// TIA Portal project "TIA1200_Level1" (V19) (continued)
REGION Network 5: Retract Cylinder B logic
   // Retract cylinder B after both cylinders are extended
   RUNG wire#powerrail
      Contact( "Gripper open" )
      Contact( "Cylinder A extended" )
      Contact( "Cylinder B extended" )
      S_SR(operand := "Retract cylinder B", r1 := wire#w1)
   END_RUNG
   RUNG wire#powerrail
      Contact( "Cylinder B retracted" )
   END_RUNG wire#w1
   // the same network as SCL:
   IF "Gripper open" AND "Cylinder A extended" AND "Cylinder B extended" THEN
       "Retract cylinder B" := TRUE;   // SR flip-flop
   END_IF;
   IF "Cylinder B retracted" THEN "Retract cylinder B" := FALSE; END_IF;
END_REGION

REGION Network 6: Retract Cylinder A Logic
   // Retract cylinder A when cylinder A is extended, cylinder B is retracted and gripper is open; stop after its upper limit
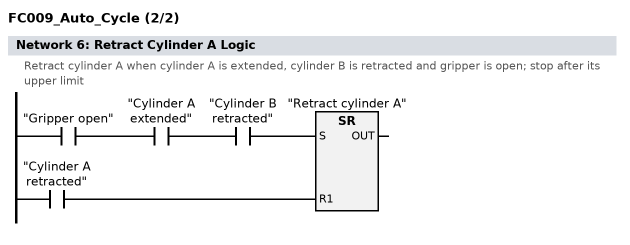
   RUNG wire#powerrail
      Contact( "Gripper open" )
      Contact( "Cylinder A extended" )
      Contact( "Cylinder B retracted" )
      S_SR(operand := "Retract cylinder A", r1 := wire#w1)
   END_RUNG
   RUNG wire#powerrail
      Contact( "Cylinder A retracted" )
   END_RUNG wire#w1
   // the same network as SCL:
   IF "Gripper open" AND "Cylinder A extended" AND "Cylinder B retracted" THEN
       "Retract cylinder A" := TRUE;   // SR flip-flop
   END_IF;
   IF "Cylinder A retracted" THEN "Retract cylinder A" := FALSE; END_IF;
END_REGION
END_FUNCTION

FUNCTION "FC010_OneButton_OneLight" : Void   // FC14, LAD
{ S7_Optimized_Access := 'TRUE' }
VERSION : 0.1
   VAR_TEMP   // added for the SCL form of the ladder/FBD networks
      _w1 : Bool;
   END_VAR
BEGIN

REGION Network 1 (FBD): Lamp Toggle Logic
   // XOR outputs 1 only when both inputs have different states; identical states produce 0
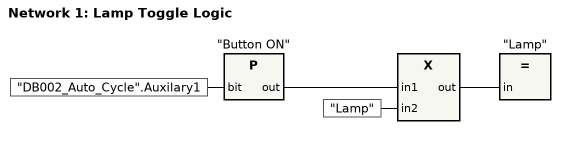
   #_w1 := "Button ON" AND NOT "DB002_Auto_Cycle".Auxilary1;   // rising edge of "Button ON"
   "DB002_Auto_Cycle".Auxilary1 := "Button ON";
   "Lamp" := #_w1 XOR "Lamp";
END_REGION
END_FUNCTION

FUNCTION "FC011_Voltage_Control" : Void   // FC15, LAD
{ S7_Optimized_Access := 'TRUE' }
VERSION : 0.1
BEGIN

REGION Network 1: Voltage Output Control Logic
   // Set QW80 to 0 V, 5 V, or 10 V depending on input states I1.0 and I1.1 (Integer range: 0 - 27648)
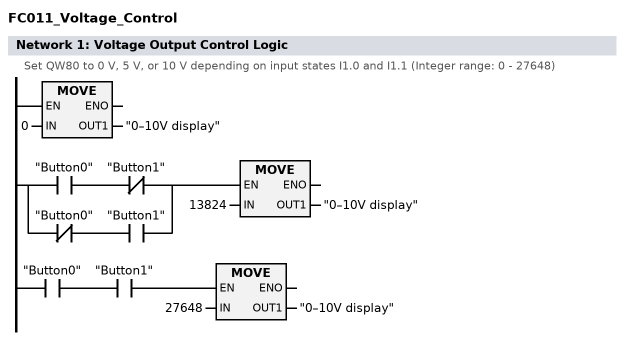
   RUNG wire#powerrail
      Move(in := 0, out1 => "0–10V display")
   END_RUNG
   RUNG wire#powerrail
      Contact( "Button0" )
      I_Contact( "Button1" )
      wire#w1
      Move(in := 13824, out1 => "0–10V display")
   END_RUNG
   RUNG wire#powerrail
      I_Contact( "Button0" )
      Contact( "Button1" )
   END_RUNG wire#w1
   RUNG wire#powerrail
      Contact( "Button0" )
      Contact( "Button1" )
      Move(in := 27648, out1 => "0–10V display")
   END_RUNG
   // the same network as SCL:
   "0–10V display" := 0;
   IF ("Button0" AND NOT "Button1") OR (NOT "Button0" AND "Button1") THEN "0–10V display" := 13824; END_IF;
   IF "Button0" AND "Button1" THEN "0–10V display" := 27648; END_IF;
END_REGION
END_FUNCTION

FUNCTION "FC012_Calculations" : Void   // FC16, LAD
{ S7_Optimized_Access := 'TRUE' }
VERSION : 0.1
   VAR_TEMP   // added for the SCL form of the ladder/FBD networks
      _w1 : Bool;
   END_VAR
BEGIN

REGION Network 1: Production Stock Calculation
   // Calculate stock = Sum1 + Sum2 − Losses
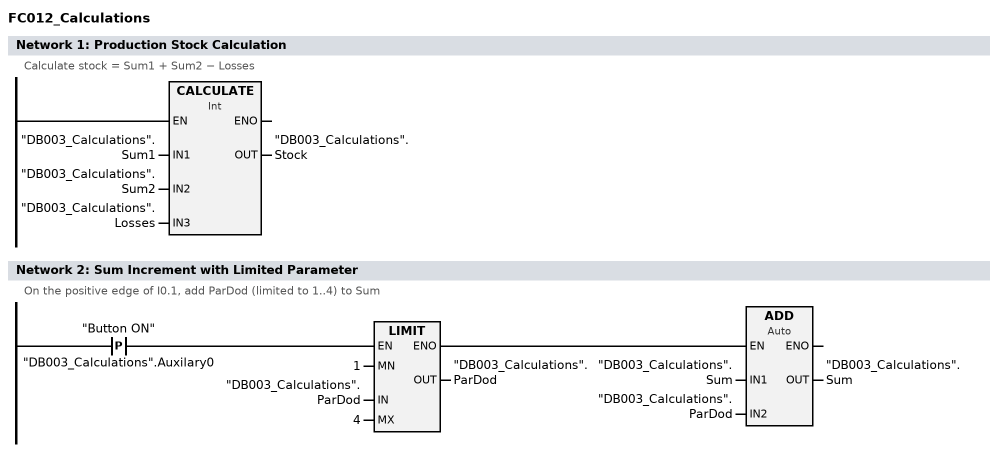
   RUNG wire#powerrail
      { S7_Templates := "SrcType := Int"; S7_Expression := "IN1 + IN2 - IN3" } Calculate(in1 := "DB003_Calculations".Sum1, in2 := "DB003_Calculations".Sum2, in3 := "DB003_Calculations".Losses, out => "DB003_Calculations".Stock)
   END_RUNG
   // the same network as SCL:
   "DB003_Calculations".Stock := "DB003_Calculations".Sum1 + "DB003_Calculations".Sum2 - "DB003_Calculations".Losses;
END_REGION

REGION Network 2: Sum Increment with Limited Parameter
   // On the positive edge of I0.1, add ParDod (limited to 1..4) to Sum
   #_w1 := "Button ON" AND NOT "DB003_Calculations".Auxilary0;   // rising edge of "Button ON"
   "DB003_Calculations".Auxilary0 := "Button ON";
   IF #_w1 THEN
       "DB003_Calculations".ParDod := LIMIT(MN := 1, IN := "DB003_Calculations".ParDod, MX := 4);
       "DB003_Calculations".Sum := "DB003_Calculations".Sum + "DB003_Calculations".ParDod;
   END_IF;
END_REGION
END_FUNCTION

FUNCTION "FC013_Labeler_Control" : Void   // FC17, LAD
{ S7_Optimized_Access := 'TRUE' }
VERSION : 0.1
   VAR_TEMP   // added for the SCL form of the ladder/FBD networks
      _w1 : Bool;
   END_VAR
BEGIN

REGION Network 1: Roll Initialization & Roll Counter
   // On Button0 load a new labels roll and increment labels roll total counter
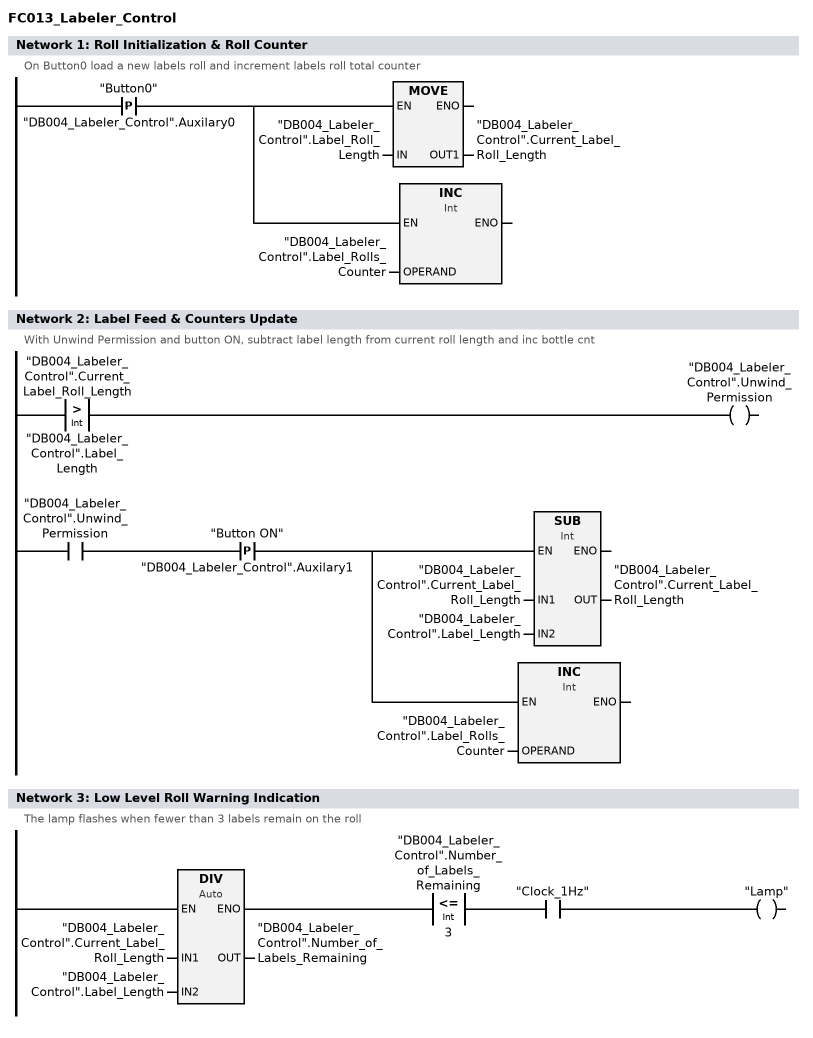
   RUNG wire#powerrail
      P_Contact(operand := "Button0", bit := "DB004_Labeler_Control".Auxilary0)
      wire#w1
      Move(in := "DB004_Labeler_Control".Label_Roll_Length, out1 => "DB004_Labeler_Control".Current_Label_Roll_Length)
   END_RUNG
   RUNG wire#w1
      { S7_Templates := "DestType := Int" } Inc( "DB004_Labeler_Control".Label_Rolls_Counter )
   END_RUNG
   // the same network as SCL:
   #_w1 := "Button0" AND NOT "DB004_Labeler_Control".Auxilary0;   // rising edge of "Button0"
   "DB004_Labeler_Control".Auxilary0 := "Button0";
   IF #_w1 THEN
       "DB004_Labeler_Control".Current_Label_Roll_Length := "DB004_Labeler_Control".Label_Roll_Length;
       "DB004_Labeler_Control".Label_Rolls_Counter := "DB004_Labeler_Control".Label_Rolls_Counter + 1;
   END_IF;
END_REGION

REGION Network 2: Label Feed & Counters Update
   // With Unwind Permission and button ON, subtract label length from current roll length and inc bottle cnt
   RUNG wire#powerrail
      { S7_Templates := "SrcType := Int" } GT_Contact(in1 := "DB004_Labeler_Control".Current_Label_Roll_Length, in2 := "DB004_Labeler_Control".Label_Length)
      Coil( "DB004_Labeler_Control".Unwind_Permission )
   END_RUNG
   RUNG wire#powerrail
      Contact( "DB004_Labeler_Control".Unwind_Permission )
      P_Contact(operand := "Button ON", bit := "DB004_Labeler_Control".Auxilary1)
      wire#w1
      { S7_Templates := "SrcType := Int" } Sub(in1 := "DB004_Labeler_Control".Current_Label_Roll_Length, in2 := "DB004_Labeler_Control".Label_Length, out => "DB004_Labeler_Control".Current_Label_Roll_Length)
   END_RUNG
   RUNG wire#w1
      { S7_Templates := "DestType := Int" } Inc( "DB004_Labeler_Control".Label_Rolls_Counter )
   END_RUNG
   // the same network as SCL:
   "DB004_Labeler_Control".Unwind_Permission := "DB004_Labeler_Control".Current_Label_Roll_Length > "DB004_Labeler_Control".Label_Length;
   #_w1 := "DB004_Labeler_Control".Unwind_Permission AND "Button ON" AND NOT "DB004_Labeler_Control".Auxilary1;   // rising edge of "Button ON"
   "DB004_Labeler_Control".Auxilary1 := "Button ON";
   IF #_w1 THEN
       "DB004_Labeler_Control".Current_Label_Roll_Length := "DB004_Labeler_Control".Current_Label_Roll_Length - "DB004_Labeler_Control".Label_Length;
       "DB004_Labeler_Control".Label_Rolls_Counter := "DB004_Labeler_Control".Label_Rolls_Counter + 1;
   END_IF;
END_REGION

REGION Network 3: Low Level Roll Warning Indication
   // The lamp flashes when fewer than 3 labels remain on the roll
   RUNG wire#powerrail
      Div(in1 := "DB004_Labeler_Control".Current_Label_Roll_Length, in2 := "DB004_Labeler_Control".Label_Length, out => "DB004_Labeler_Control".Number_of_Labels_Remaining)
      { S7_Templates := "SrcType := Int" } LE_Contact(in1 := "DB004_Labeler_Control".Number_of_Labels_Remaining, in2 := 3)
      Contact( "Clock_1Hz" )
      Coil( "Lamp" )
   END_RUNG
   // the same network as SCL:
   "DB004_Labeler_Control".Number_of_Labels_Remaining := "DB004_Labeler_Control".Current_Label_Roll_Length / "DB004_Labeler_Control".Label_Length;
   "Lamp" := ("DB004_Labeler_Control".Number_of_Labels_Remaining <= 3) AND "Clock_1Hz";
END_REGION
END_FUNCTION

FUNCTION "FC014_Buffer_Filling" : Void   // FC18, LAD
{ S7_Optimized_Access := 'TRUE' }
VERSION : 0.1
BEGIN

REGION Network 1: Buffer Counter & Limits Logic
   // Count up on I1.3 and down on I1.5 with CTUD (PV=10). NOT QU blocks further up-counting at full; reset with I0.0
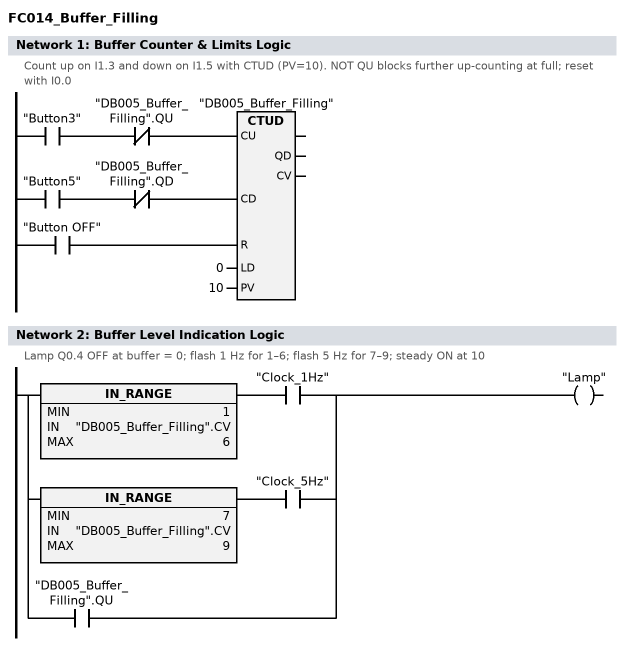
   "DB005_Buffer_Filling".CTUD(CU := "Button3" AND NOT "DB005_Buffer_Filling".QU,
                           CD := "Button5" AND NOT "DB005_Buffer_Filling".QD,
                           R := "Button OFF",
                           LD := 0,
                           PV := 10);
END_REGION

REGION Network 2: Buffer Level Indication Logic
   // Lamp Q0.4 OFF at buffer = 0; flash 1 Hz for 1–6; flash 5 Hz for 7–9; steady ON at 10
   RUNG wire#powerrail
      { S7_Templates := "SrcType := Int" } InRange(min := 1, in := "DB005_Buffer_Filling".CV, max := 6)
      Contact( "Clock_1Hz" )
      wire#w1
      Coil( "Lamp" )
   END_RUNG
   RUNG wire#powerrail
      { S7_Templates := "SrcType := Int" } InRange(min := 7, in := "DB005_Buffer_Filling".CV, max := 9)
      Contact( "Clock_5Hz" )
   END_RUNG wire#w1
   RUNG wire#powerrail
      Contact( "DB005_Buffer_Filling".QU )
   END_RUNG wire#w1
   // the same network as SCL:
   "Lamp" := ((1 <= "DB005_Buffer_Filling".CV) AND ("DB005_Buffer_Filling".CV <= 6) AND "Clock_1Hz") OR ((7 <= "DB005_Buffer_Filling".CV) AND ("DB005_Buffer_Filling".CV <= 9) AND "Clock_5Hz") OR "DB005_Buffer_Filling".QU;
END_REGION
END_FUNCTION

FUNCTION "FC015_Lift_Sequence" : Void   // FC19, LAD
{ S7_Optimized_Access := 'TRUE' }
VERSION : 0.1
BEGIN

REGION Network 1: Sequence Step Counter Logic
   // On the positive edge of I0.1, increment the step counter; use CTU for steps 1..13
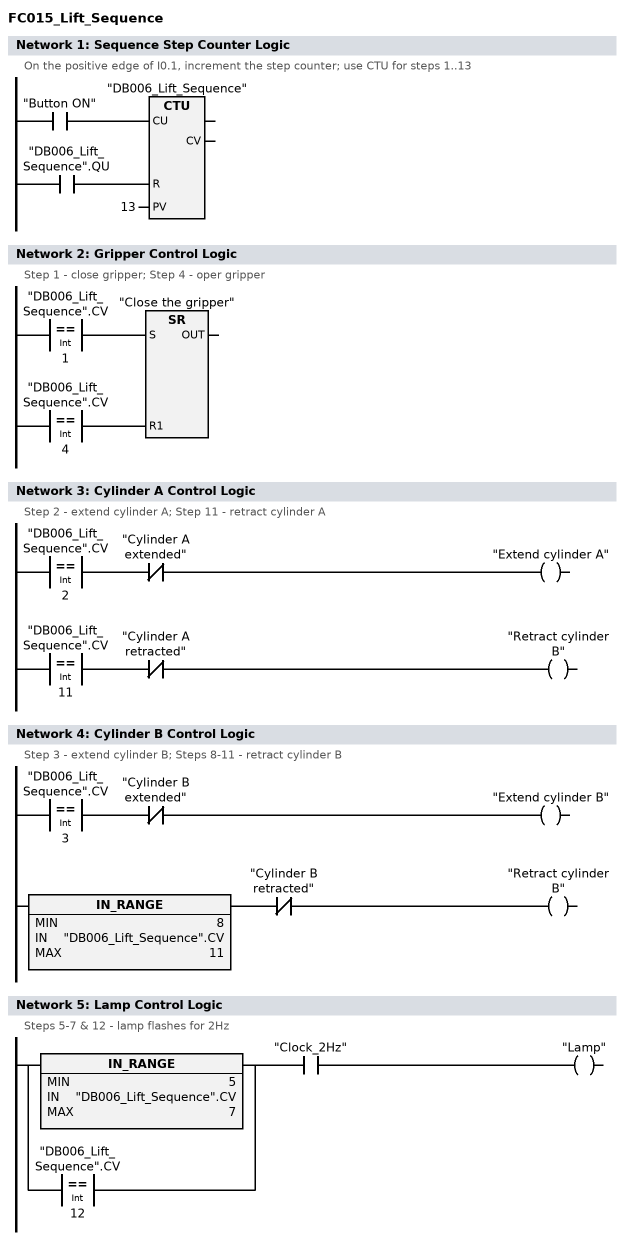
   "DB006_Lift_Sequence".CTU(CU := "Button ON", R := "DB006_Lift_Sequence".QU, PV := 13);
END_REGION

REGION Network 2: Gripper Control Logic
   // Step 1 - close gripper; Step 4 - oper gripper
   RUNG wire#powerrail
      { S7_Templates := "SrcType := Int" } EQ_Contact(in1 := "DB006_Lift_Sequence".CV, in2 := 1)
      S_SR(operand := "Close the gripper", r1 := wire#w1)
   END_RUNG
   RUNG wire#powerrail
      { S7_Templates := "SrcType := Int" } EQ_Contact(in1 := "DB006_Lift_Sequence".CV, in2 := 4)
   END_RUNG wire#w1
   // the same network as SCL:
   IF "DB006_Lift_Sequence".CV = 1 THEN
       "Close the gripper" := TRUE;   // SR flip-flop
   END_IF;
   IF "DB006_Lift_Sequence".CV = 4 THEN "Close the gripper" := FALSE; END_IF;
END_REGION

REGION Network 3: Cylinder A Control Logic
   // Step 2 - extend cylinder A; Step 11 - retract cylinder A
   RUNG wire#powerrail
      { S7_Templates := "SrcType := Int" } EQ_Contact(in1 := "DB006_Lift_Sequence".CV, in2 := 2)
      I_Contact( "Cylinder A extended" )
      Coil( "Extend cylinder A" )
   END_RUNG
   RUNG wire#powerrail
      { S7_Templates := "SrcType := Int" } EQ_Contact(in1 := "DB006_Lift_Sequence".CV, in2 := 11)
      I_Contact( "Cylinder A retracted" )
      Coil( "Retract cylinder B" )
   END_RUNG
   // the same network as SCL:
   "Extend cylinder A" := ("DB006_Lift_Sequence".CV = 2) AND NOT "Cylinder A extended";
   "Retract cylinder B" := ("DB006_Lift_Sequence".CV = 11) AND NOT "Cylinder A retracted";
END_REGION

REGION Network 4: Cylinder B Control Logic
   // Step 3 - extend cylinder B; Steps 8-11 - retract cylinder B
   RUNG wire#powerrail
      { S7_Templates := "SrcType := Int" } EQ_Contact(in1 := "DB006_Lift_Sequence".CV, in2 := 3)
      I_Contact( "Cylinder B extended" )
      Coil( "Extend cylinder B" )
   END_RUNG
   RUNG wire#powerrail
      { S7_Templates := "SrcType := Int" } InRange(min := 8, in := "DB006_Lift_Sequence".CV, max := 11)
      I_Contact( "Cylinder B retracted" )
      Coil( "Retract cylinder B" )
   END_RUNG
   // the same network as SCL:
   "Extend cylinder B" := ("DB006_Lift_Sequence".CV = 3) AND NOT "Cylinder B extended";
   "Retract cylinder B" := (8 <= "DB006_Lift_Sequence".CV) AND ("DB006_Lift_Sequence".CV <= 11) AND NOT "Cylinder B retracted";
END_REGION

REGION Network 5: Lamp Control Logic
   // Steps 5-7 & 12 - lamp flashes for 2Hz
   RUNG wire#powerrail
      { S7_Templates := "SrcType := Int" } InRange(min := 5, in := "DB006_Lift_Sequence".CV, max := 7)
      wire#w1
      Contact( "Clock_2Hz" )
      Coil( "Lamp" )
   END_RUNG
   RUNG wire#powerrail
      { S7_Templates := "SrcType := Int" } EQ_Contact(in1 := "DB006_Lift_Sequence".CV, in2 := 12)
   END_RUNG wire#w1
   // the same network as SCL:
   "Lamp" := (((5 <= "DB006_Lift_Sequence".CV) AND ("DB006_Lift_Sequence".CV <= 7)) OR ("DB006_Lift_Sequence".CV = 12)) AND "Clock_2Hz";
END_REGION
END_FUNCTION

FUNCTION "FC016_Pulse_Generator" : Void   // FC20, LAD
{ S7_Optimized_Access := 'TRUE' }
VERSION : 0.1
BEGIN

REGION Network 1: Pulse Generator Enable Logic
   // Button I0.1 starts the pulse generator; I0.0 stops it
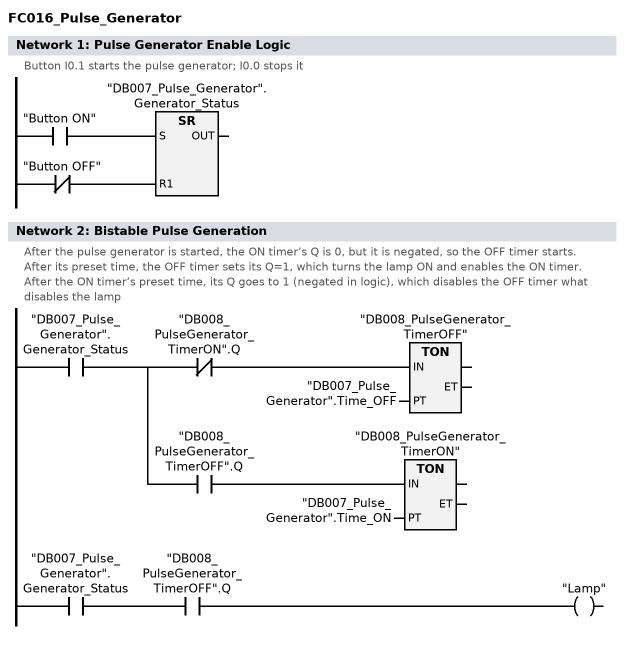
   RUNG wire#powerrail
      Contact( "Button ON" )
      S_SR(operand := "DB007_Pulse_Generator".Generator_Status, r1 := wire#w1)
   END_RUNG
   RUNG wire#powerrail
      I_Contact( "Button OFF" )
   END_RUNG wire#w1
   // the same network as SCL:
   IF "Button ON" THEN
       "DB007_Pulse_Generator".Generator_Status := TRUE;   // SR flip-flop
   END_IF;
   IF NOT "Button OFF" THEN "DB007_Pulse_Generator".Generator_Status := FALSE; END_IF;
END_REGION

REGION Network 2: Bistable Pulse Generation
   // After the pulse generator is started, the ON timer’s Q is 0, but it is negated, so the OFF timer starts. 
   // After its preset time, the OFF timer sets its Q=1, which turns the lamp ON and enables the ON timer. 
   // After the ON timer’s preset time, its Q goes to 1 (negated in logic), which disables the OFF timer what disables the lamp
   "DB008_PulseGenerator_TimerOFF".TON(IN := "DB007_Pulse_Generator".Generator_Status AND NOT "DB008_PulseGenerator_TimerON".Q,
                           PT := "DB007_Pulse_Generator".Time_OFF);
   "DB008_PulseGenerator_TimerON".TON(IN := "DB007_Pulse_Generator".Generator_Status AND "DB008_PulseGenerator_TimerOFF".Q,
                           PT := "DB007_Pulse_Generator".Time_ON);
   "Lamp" := "DB007_Pulse_Generator".Generator_Status AND "DB008_PulseGenerator_TimerOFF".Q;
END_REGION
END_FUNCTION

FUNCTION "FC017_Motor_With_Cooling" : Void   // FC21, LAD
{ S7_Optimized_Access := 'TRUE' }
VERSION : 0.1
   VAR_TEMP   // added for the SCL form of the ladder/FBD networks
      _w1 : Bool;
   END_VAR
BEGIN

REGION Network 1: E‑Stop Alarm & Immediate Stop
   // E‑Stop I0.2 instantly stops motor and fan and latches "E-Stop Alarm"; reset the alarm with I1.5
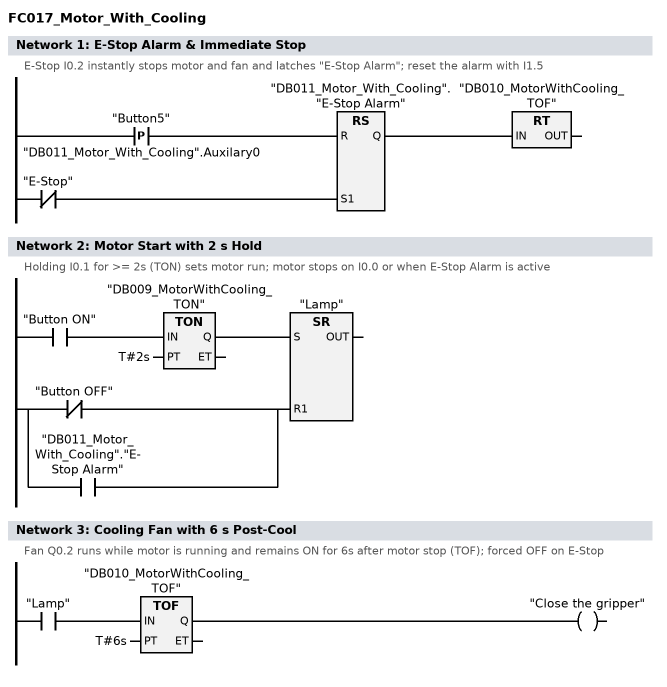
   RUNG wire#powerrail
      P_Contact(operand := "Button5", bit := "DB011_Motor_With_Cooling".Auxilary0)
      S_RS(operand := "DB011_Motor_With_Cooling"."E-Stop Alarm", s1 := wire#w1)
      RT_Coil( "DB010_MotorWithCooling_TOF" )
   END_RUNG
   RUNG wire#powerrail
      I_Contact( "E-Stop" )
   END_RUNG wire#w1
   // the same network as SCL:
   #_w1 := "Button5" AND NOT "DB011_Motor_With_Cooling".Auxilary0;   // rising edge of "Button5"
   "DB011_Motor_With_Cooling".Auxilary0 := "Button5";
   IF #_w1 THEN
       "DB011_Motor_With_Cooling"."E-Stop Alarm" := FALSE;   // RS flip-flop
   END_IF;
   IF NOT "E-Stop" THEN "DB011_Motor_With_Cooling"."E-Stop Alarm" := TRUE; END_IF;
   IF "DB011_Motor_With_Cooling"."E-Stop Alarm" THEN RESET_TIMER("DB010_MotorWithCooling_TOF"); END_IF;
END_REGION

REGION Network 2: Motor Start with 2 s Hold
   // Holding I0.1 for >= 2s (TON) sets motor run; motor stops on I0.0 or when E-Stop Alarm is active
   "DB009_MotorWithCooling_TON".TON(IN := "Button ON", PT := T#2s);
   IF "DB009_MotorWithCooling_TON".Q THEN
       "Lamp" := TRUE;   // SR flip-flop
   END_IF;
   IF NOT "Button OFF" OR "DB011_Motor_With_Cooling"."E-Stop Alarm" THEN "Lamp" := FALSE; END_IF;
END_REGION

REGION Network 3: Cooling Fan with 6 s Post‑Cool
   // Fan Q0.2 runs while motor is running and remains ON for 6s after motor stop (TOF); forced OFF on E‑Stop
   "DB010_MotorWithCooling_TOF".TOF(IN := "Lamp", PT := T#6s);
   "Close the gripper" := "DB010_MotorWithCooling_TOF".Q;
END_REGION
END_FUNCTION

FUNCTION "FC018_Cylinder_Timeout" : Void   // FC22, LAD
{ S7_Optimized_Access := 'TRUE' }
VERSION : 0.1
   VAR_TEMP   // added for the SCL form of the ladder/FBD networks
      _w1 : Bool;
   END_VAR
BEGIN

REGION Network 1: Motion Timeout Detection & Alarm Set
   // If cylinder moves for >= 2 s without reaching the target sensor, set Timeout Alarm. Reset the alarm with I1.5; blink lamp Q0.4 at 1 Hz when the alarm is active
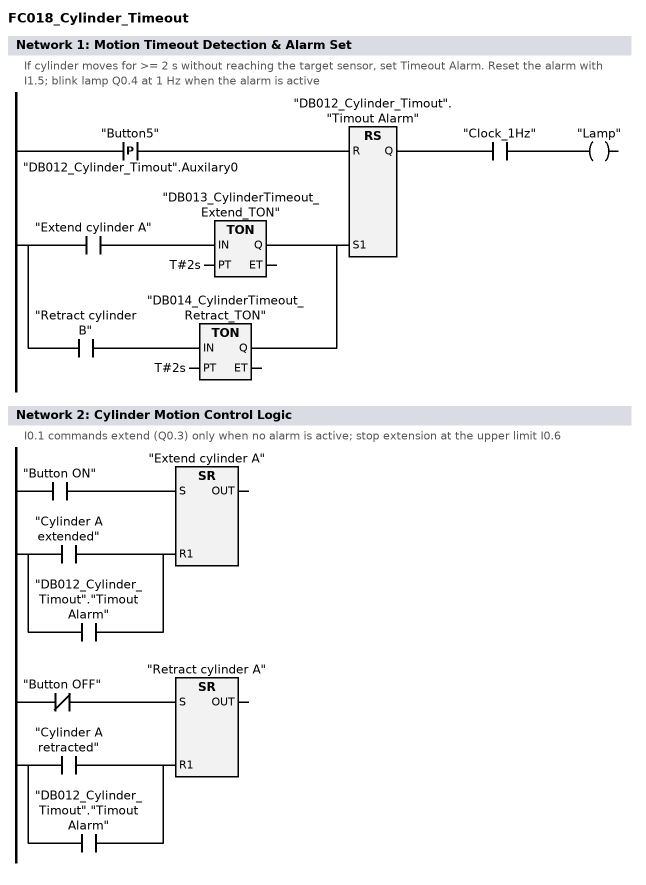
   #_w1 := "Button5" AND NOT "DB012_Cylinder_Timout".Auxilary0;   // rising edge of "Button5"
   "DB012_Cylinder_Timout".Auxilary0 := "Button5";
   "DB013_CylinderTimeout_Extend_TON".TON(IN := "Extend cylinder A", PT := T#2s);
   "DB014_CylinderTimeout_Retract_TON".TON(IN := "Retract cylinder B", PT := T#2s);
   IF #_w1 THEN
       "DB012_Cylinder_Timout"."Timout Alarm" := FALSE;   // RS flip-flop
   END_IF;
   IF "DB013_CylinderTimeout_Extend_TON".Q OR "DB014_CylinderTimeout_Retract_TON".Q THEN
       "DB012_Cylinder_Timout"."Timout Alarm" := TRUE;
   END_IF;
   "Lamp" := "DB012_Cylinder_Timout"."Timout Alarm" AND "Clock_1Hz";
END_REGION

REGION Network 2: Cylinder Motion Control Logic
   // I0.1 commands extend (Q0.3) only when no alarm is active; stop extension at the upper limit I0.6
   RUNG wire#powerrail
      Contact( "Button ON" )
      S_SR(operand := "Extend cylinder A", r1 := wire#w1)
   END_RUNG
   RUNG wire#powerrail
      Contact( "Cylinder A extended" )
   END_RUNG wire#w1
   RUNG wire#powerrail
      Contact( "DB012_Cylinder_Timout"."Timout Alarm" )
   END_RUNG wire#w1
   RUNG wire#powerrail
      I_Contact( "Button OFF" )
      S_SR(operand := "Retract cylinder A", r1 := wire#w2)
   END_RUNG
   RUNG wire#powerrail
      Contact( "Cylinder A retracted" )
   END_RUNG wire#w2
   RUNG wire#powerrail
      Contact( "DB012_Cylinder_Timout"."Timout Alarm" )
   END_RUNG wire#w2
   // the same network as SCL:
   IF "Button ON" THEN
       "Extend cylinder A" := TRUE;   // SR flip-flop
   END_IF;
   IF "Cylinder A extended" OR "DB012_Cylinder_Timout"."Timout Alarm" THEN
       "Extend cylinder A" := FALSE;
   END_IF;
   IF NOT "Button OFF" THEN
       "Retract cylinder A" := TRUE;   // SR flip-flop
   END_IF;
   IF "Cylinder A retracted" OR "DB012_Cylinder_Timout"."Timout Alarm" THEN
       "Retract cylinder A" := FALSE;
   END_IF;
END_REGION
END_FUNCTION

FUNCTION "FC004_EndPosition#2" : Void   // FC23, LAD
{ S7_Optimized_Access := 'TRUE' }
VERSION : 0.1
BEGIN

REGION Network 1: Extend Cylinder A Logic
   // Button ON extends cylinder A until the upper limit I0.6 is reached
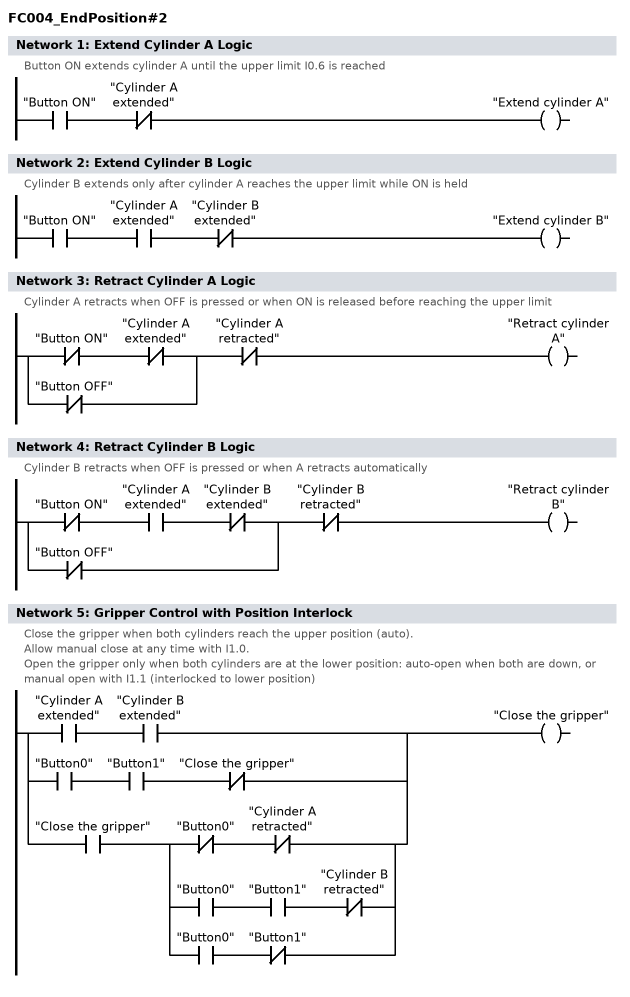
   RUNG wire#powerrail
      Contact( "Button ON" )
      I_Contact( "Cylinder A extended" )
      Coil( "Extend cylinder A" )
   END_RUNG
   // the same network as SCL:
   "Extend cylinder A" := "Button ON" AND NOT "Cylinder A extended";
END_REGION

REGION Network 2: Extend Cylinder B Logic
   // Cylinder B extends only after cylinder A reaches the upper limit while ON is held
   RUNG wire#powerrail
      Contact( "Button ON" )
      Contact( "Cylinder A extended" )
      I_Contact( "Cylinder B extended" )
      Coil( "Extend cylinder B" )
   END_RUNG
   // the same network as SCL:
   "Extend cylinder B" := "Button ON" AND "Cylinder A extended" AND NOT "Cylinder B extended";
END_REGION

REGION Network 3: Retract Cylinder A Logic
   // Cylinder A retracts when OFF is pressed or when ON is released before reaching the upper limit
   RUNG wire#powerrail
      I_Contact( "Button ON" )
      I_Contact( "Cylinder A extended" )
      wire#w1
      I_Contact( "Cylinder A retracted" )
      Coil( "Retract cylinder A" )
   END_RUNG
   RUNG wire#powerrail
      I_Contact( "Button OFF" )
   END_RUNG wire#w1
   // the same network as SCL:
   "Retract cylinder A" := ((NOT "Button ON" AND NOT "Cylinder A extended") OR NOT "Button OFF") AND NOT "Cylinder A retracted";
END_REGION

REGION Network 4: Retract Cylinder B Logic
   // Cylinder B retracts when OFF is pressed or when A retracts automatically
   RUNG wire#powerrail
      I_Contact( "Button ON" )
      Contact( "Cylinder A extended" )
      I_Contact( "Cylinder B extended" )
      wire#w1
      I_Contact( "Cylinder B retracted" )
      Coil( "Retract cylinder B" )
   END_RUNG
   RUNG wire#powerrail
      I_Contact( "Button OFF" )
   END_RUNG wire#w1
   // the same network as SCL:
   "Retract cylinder B" := ((NOT "Button ON" AND "Cylinder A extended" AND NOT "Cylinder B extended") OR NOT "Button OFF") AND NOT "Cylinder B retracted";
END_REGION

REGION Network 5: Gripper Control with Position Interlock
   // Close the gripper when both cylinders reach the upper position (auto). 
   // Allow manual close at any time with I1.0. 
   // Open the gripper only when both cylinders are at the lower position: auto‑open when both are down, or manual open with I1.1 (interlocked to lower position)
   RUNG wire#powerrail
      Contact( "Cylinder A extended" )
      Contact( "Cylinder B extended" )
      wire#w1
      Coil( "Close the gripper" )
   END_RUNG
   RUNG wire#powerrail
      Contact( "Button0" )
      Contact( "Button1" )
      I_Contact( "Close the gripper" )
   END_RUNG wire#w1
   RUNG wire#powerrail
      Contact( "Close the gripper" )
      wire#w2
      I_Contact( "Button0" )
      I_Contact( "Cylinder A retracted" )
   END_RUNG wire#w1
   RUNG wire#w2
      Contact( "Button0" )
      Contact( "Button1" )
      I_Contact( "Cylinder B retracted" )
   END_RUNG wire#w1
   RUNG wire#w2
      Contact( "Button0" )
      I_Contact( "Button1" )
   END_RUNG wire#w1
   // the same network as SCL:
   "Close the gripper" := ("Cylinder A extended" AND "Cylinder B extended") OR ("Button0" AND "Button1" AND NOT "Close the gripper") OR ("Close the gripper" AND ((NOT "Button0" AND NOT "Cylinder A retracted") OR ("Button0" AND "Button1" AND NOT "Cylinder B retracted") OR ("Button0" AND NOT "Button1")));
END_REGION
END_FUNCTION

FUNCTION "FC019_Manual_Sequence" : Void   // FC24, FBD
{ S7_Optimized_Access := 'TRUE' }
VERSION : 0.1
BEGIN

REGION Network 1: Manual Sequence Step#1
   // Pressing button I1.0 extends cylinder A and turns the lamp ON
